           IF #Request AND NOT "PN_Mixinghead".Mixinghead[#MH].ReinigungskolbenDigital.ChckConnFault THEN
               "PN_Mixinghead".Mixinghead[#MH].ReinigungskolbenDigital.GeneralParameters.Request := "PN_Mixinghead".Mixinghead[#MH].ReinigungskolbenDigital.Active;
               "PN_Mixinghead".Mixinghead[#MH].ReinigungskolbenDigital.Zeiten.Request := "PN_Mixinghead".Mixinghead[#MH].ReinigungskolbenDigital.Active;
           END_IF;

           "WRREC_FC"(GOON := #GOON,
                      REQ := "PN_Mixinghead".Mixinghead[#MH].ReinigungskolbenDigital.GeneralParameters.Request,
                      ADDRESS := #TempHWID,
                      INDEX := #IDM_CleaningPiston_Digital_GeneralParameters_Index,
                      LENGTH := #IDM_CleaningPiston_Digital_GeneralParameters_Length,
                      WRREC_DONE => #t.DONE,
                      WRREC_BUSY => #t.BUSY,
                      WRREC_ERROR => #t.ERROR,
                      WRREC_STATUS => #t.STATUS,
                      ACTIVE := "PN_Mixinghead".Mixinghead[#MH].ReinigungskolbenDigital.Active,
                      RECORD := "PN_Mixinghead".Mixinghead[#MH].ReinigungskolbenDigital.GeneralParameters.Data,
                      DONE := "PN_Mixinghead".Mixinghead[#MH].ReinigungskolbenDigital.GeneralParameters.Transmitting);

           "WRREC_FC"(GOON := #GOON,
                      REQ := "PN_Mixinghead".Mixinghead[#MH].ReinigungskolbenDigital.Zeiten.Request,
                      ADDRESS := #TempHWID,
                      INDEX := #IDM_CleaningPiston_Digital_Zeiten_Index,
                      LENGTH := #IDM_CleaningPiston_Digital_Zeiten_Length,
                      WRREC_DONE => #t.DONE,
                      WRREC_BUSY => #t.BUSY,
                      WRREC_ERROR => #t.ERROR,
                      WRREC_STATUS => #t.STATUS,
                      ACTIVE := "PN_Mixinghead".Mixinghead[#MH].ReinigungskolbenDigital.Active,
                      RECORD := "PN_Mixinghead".Mixinghead[#MH].ReinigungskolbenDigital.Zeiten.Data,
                      DONE := "PN_Mixinghead".Mixinghead[#MH].ReinigungskolbenDigital.Zeiten.Transmitting);
       END_IF;

       // -----------------------------------
       // REINIGUNGSKOLBEN geregelt   
       // -----------------------------------
       IF "PN_Mixinghead".Mixinghead[#MH].ReinigungskolbenGeregelt.Active THEN
           #Address := INT_TO_WORD("PN_Mixinghead".Mixinghead[#MH].ReinigungskolbenGeregelt.Address);
           #ReturnValue := LOG2MOD(IOID := B#16#54, ADDR := #Address, HWID => #TempHWID);
           // Kommunikationsüberwachung
           // Nach einem Verbindungsabbruch werden die Telegramme automatisch verschickt.
           #Request := false;
           "CHCKPNCONN"(GOON := #GOON,
                        Active := "PN_Mixinghead".Mixinghead[#MH].ReinigungskolbenGeregelt.Active,
                        Address := #TempHWID,
                        PN_Request := #Request,
                        PN_Fault := "PN_Mixinghead".Mixinghead[#MH].ReinigungskolbenGeregelt.ChckConnFault,
                        DONE := "PN_Mixinghead".Mixinghead[#MH].ReinigungskolbenGeregelt.ChckConnDone);

           IF #Request AND NOT "PN_Mixinghead".Mixinghead[#MH].ReinigungskolbenGeregelt.ChckConnFault THEN
               "PN_Mixinghead".Mixinghead[#MH].ReinigungskolbenGeregelt.GeneralParameters.Request := "PN_Mixinghead".Mixinghead[#MH].ReinigungskolbenGeregelt.Active;
               "PN_Mixinghead".Mixinghead[#MH].ReinigungskolbenGeregelt.Zeiten.Request := "PN_Mixinghead".Mixinghead[#MH].ReinigungskolbenGeregelt.Active;
               "PN_Mixinghead".Mixinghead[#MH].ReinigungskolbenGeregelt.Skalierung.Request := "PN_Mixinghead".Mixinghead[#MH].ReinigungskolbenGeregelt.Active;
               "PN_Mixinghead".Mixinghead[#MH].ReinigungskolbenGeregelt.Regelparameter.Request := "PN_Mixinghead".Mixinghead[#MH].ReinigungskolbenGeregelt.Active;
           END_IF;

           "WRREC_FC"(GOON := #GOON,
                      REQ := "PN_Mixinghead".Mixinghead[#MH].ReinigungskolbenGeregelt.GeneralParameters.Request,
                      ACTIVE := "PN_Mixinghead".Mixinghead[#MH].ReinigungskolbenGeregelt.Active,
                      ADDRESS := #TempHWID,
                      INDEX := #IDM_CleaningPiston_Analog_Loop_GeneralParameters_Index,
                      LENGTH := #IDM_CleaningPiston_Analog_Loop_GeneralParameters_Length,
                      WRREC_DONE => #t.DONE,
                      WRREC_BUSY => #t.BUSY,
                      WRREC_ERROR => #t.ERROR,
                      WRREC_STATUS => #t.STATUS,
                      RECORD := "PN_Mixinghead".Mixinghead[#MH].ReinigungskolbenGeregelt.GeneralParameters.Data,
                      DONE := "PN_Mixinghead".Mixinghead[#MH].ReinigungskolbenGeregelt.GeneralParameters.Transmitting);

           "WRREC_FC"(GOON := #GOON,
                      REQ := "PN_Mixinghead".Mixinghead[#MH].ReinigungskolbenGeregelt.Zeiten.Request,
                      ACTIVE := "PN_Mixinghead".Mixinghead[#MH].ReinigungskolbenGeregelt.Active,
                      ADDRESS := #TempHWID,
                      INDEX := #IDM_CleaningPiston_Analog_Loop_Zeiten_Index,
                      LENGTH := #IDM_CleaningPiston_Analog_Loop_Zeiten_Length,
                      WRREC_DONE => #t.DONE,
                      WRREC_BUSY => #t.BUSY,
                      WRREC_ERROR => #t.ERROR,
                      WRREC_STATUS => #t.STATUS,
                      RECORD := "PN_Mixinghead".Mixinghead[#MH].ReinigungskolbenGeregelt.Zeiten.Data,
                      DONE := "PN_Mixinghead".Mixinghead[#MH].ReinigungskolbenGeregelt.Zeiten.Transmitting);

           "WRREC_FC"(GOON := #GOON,
                      REQ := "PN_Mixinghead".Mixinghead[#MH].ReinigungskolbenGeregelt.Skalierung.Request,
                      ACTIVE := "PN_Mixinghead".Mixinghead[#MH].ReinigungskolbenGeregelt.Active,
                      ADDRESS := #TempHWID,
                      INDEX := #IDM_Mixinghead_Digital_GeneralParameters_Index,
                      LENGTH := #IDM_Mixinghead_Digital_GeneralParameters_Length,
                      WRREC_DONE => #t.DONE,
                      WRREC_BUSY => #t.BUSY,
                      WRREC_ERROR => #t.ERROR,
                      WRREC_STATUS => #t.STATUS,
                      RECORD := "PN_Mixinghead".Mixinghead[#MH].ReinigungskolbenGeregelt.Skalierung.Data,
                      DONE := "PN_Mixinghead".Mixinghead[#MH].ReinigungskolbenGeregelt.Skalierung.Transmitting);

           "WRREC_FC"(GOON := #GOON,
                      REQ := "PN_Mixinghead".Mixinghead[#MH].ReinigungskolbenGeregelt.Regelparameter.Request,
                      ACTIVE := "PN_Mixinghead".Mixinghead[#MH].ReinigungskolbenGeregelt.Active,
                      ADDRESS := #TempHWID,
                      INDEX := #IDM_CleaningPiston_Analog_Loop_Regelparameter_Index,
                      LENGTH := #IDM_CleaningPiston_Analog_Loop_Regelparameter_Length,
                      WRREC_DONE => #t.DONE,
                      WRREC_BUSY => #t.BUSY,
                      WRREC_ERROR => #t.ERROR,
                      WRREC_STATUS => #t.STATUS,
                      RECORD := "PN_Mixinghead".Mixinghead[#MH].ReinigungskolbenGeregelt.Regelparameter.Data,
                      DONE := "PN_Mixinghead".Mixinghead[#MH].ReinigungskolbenGeregelt.Regelparameter.Transmitting);
       END_IF;

       // -----------------------------------
       // REINIGUNGSKOLBEN gesteuert   
       // -----------------------------------
       IF "PN_Mixinghead".Mixinghead[#MH].ReinigungskolbenGesteuert.Active THEN
           #Address := INT_TO_WORD("PN_Mixinghead".Mixinghead[#MH].ReinigungskolbenGesteuert.Address);
           #ReturnValue := LOG2MOD(IOID := B#16#54, ADDR := #Address, HWID => #TempHWID);
           // Kommunikationsüberwachung
           // Nach einem Verbindungsabbruch werden die Telegramme automatisch verschickt.
           #Request := false;
           "CHCKPNCONN"(GOON := #GOON,
                        Active := "PN_Mixinghead".Mixinghead[#MH].ReinigungskolbenGesteuert.Active,
                        Address := #TempHWID,
                        PN_Request := #Request,
                        PN_Fault := "PN_Mixinghead".Mixinghead[#MH].ReinigungskolbenGesteuert.ChckConnFault,
                        DONE := "PN_Mixinghead".Mixinghead[#MH].ReinigungskolbenGesteuert.ChckConnDone);

           IF #Request AND NOT "PN_Mixinghead".Mixinghead[#MH].ReinigungskolbenGesteuert.ChckConnFault THEN
               "PN_Mixinghead".Mixinghead[#MH].ReinigungskolbenGesteuert.GeneralParameters.Request := "PN_Mixinghead".Mixinghead[#MH].ReinigungskolbenGesteuert.Active;
               "PN_Mixinghead".Mixinghead[#MH].ReinigungskolbenGesteuert.Zeiten.Request := "PN_Mixinghead".Mixinghead[#MH].ReinigungskolbenGesteuert.Active;
               "PN_Mixinghead".Mixinghead[#MH].ReinigungskolbenGesteuert.Skalierung.Request := "PN_Mixinghead".Mixinghead[#MH].ReinigungskolbenGesteuert.Active;
               "PN_Mixinghead".Mixinghead[#MH].ReinigungskolbenGesteuert.StufenAktivierung.Request := "PN_Mixinghead".Mixinghead[#MH].ReinigungskolbenGesteuert.Active;
               "PN_Mixinghead".Mixinghead[#MH].ReinigungskolbenGesteuert.StufenRückkehr.Request := "PN_Mixinghead".Mixinghead[#MH].ReinigungskolbenGesteuert.Active;
           END_IF;

           "WRREC_FC"(GOON := #GOON,
                      REQ := "PN_Mixinghead".Mixinghead[#MH].ReinigungskolbenGesteuert.GeneralParameters.Request,
                      ACTIVE := "PN_Mixinghead".Mixinghead[#MH].ReinigungskolbenGesteuert.Active,
                      ADDRESS := #TempHWID,
                      INDEX := #IDM_CleaningPiston_Analog_GeneralParameters_Index,
                      LENGTH := #IDM_CleaningPiston_Analog_GeneralParameters_Length,
                      WRREC_DONE => #t.DONE,
                      WRREC_BUSY => #t.BUSY,
                      WRREC_ERROR => #t.ERROR,
                      WRREC_STATUS => #t.STATUS,
                      RECORD := "PN_Mixinghead".Mixinghead[#MH].ReinigungskolbenGesteuert.GeneralParameters.Data,
                      DONE := "PN_Mixinghead".Mixinghead[#MH].ReinigungskolbenGesteuert.GeneralParameters.Transmitting);

           "WRREC_FC"(GOON := #GOON,
                      REQ := "PN_Mixinghead".Mixinghead[#MH].ReinigungskolbenGesteuert.Zeiten.Request,
                      ACTIVE := "PN_Mixinghead".Mixinghead[#MH].ReinigungskolbenGesteuert.Active,
                      ADDRESS := #TempHWID,
                      INDEX := #IDM_CleaningPiston_Analog_Zeiten_Index,
                      LENGTH := #IDM_CleaningPiston_Analog_Zeiten_Length,
                      WRREC_DONE => #t.DONE,
                      WRREC_BUSY => #t.BUSY,
                      WRREC_ERROR => #t.ERROR,
                      WRREC_STATUS => #t.STATUS,
                      RECORD := "PN_Mixinghead".Mixinghead[#MH].ReinigungskolbenGesteuert.Zeiten.Data,
                      DONE := "PN_Mixinghead".Mixinghead[#MH].ReinigungskolbenGesteuert.Zeiten.Transmitting);

           "WRREC_FC"(GOON := #GOON,
                      REQ := "PN_Mixinghead".Mixinghead[#MH].ReinigungskolbenGesteuert.Skalierung.Request,
                      ACTIVE := "PN_Mixinghead".Mixinghead[#MH].ReinigungskolbenGesteuert.Active,
                      ADDRESS := #TempHWID,
                      INDEX := #IDM_CleaningPiston_Analog_Skalierung_Index,
                      LENGTH := #IDM_CleaningPiston_Analog_Skalierung_Length,
                      WRREC_DONE => #t.DONE,
                      WRREC_BUSY => #t.BUSY,
                      WRREC_ERROR => #t.ERROR,
                      WRREC_STATUS => #t.STATUS,
                      RECORD := "PN_Mixinghead".Mixinghead[#MH].ReinigungskolbenGesteuert.Skalierung.Data,
                      DONE := "PN_Mixinghead".Mixinghead[#MH].ReinigungskolbenGesteuert.Skalierung.Transmitting);

           "WRREC_FC"(GOON := #GOON,
                      REQ := "PN_Mixinghead".Mixinghead[#MH].ReinigungskolbenGesteuert.StufenAktivierung.Request,
                      ACTIVE := "PN_Mixinghead".Mixinghead[#MH].ReinigungskolbenGesteuert.Active,
                      ADDRESS := #TempHWID,
                      INDEX := #IDM_CleaningPiston_Analog_StufenAktivierung_Index,
                      LENGTH := #IDM_CleaningPiston_Analog_StufenAktivierung_Length,
                      WRREC_DONE => #t.DONE,
                      WRREC_BUSY => #t.BUSY,
                      WRREC_ERROR => #t.ERROR,
                      WRREC_STATUS => #t.STATUS,
                      RECORD := "PN_Mixinghead".Mixinghead[#MH].ReinigungskolbenGesteuert.StufenAktivierung.Data,
                      DONE := "PN_Mixinghead".Mixinghead[#MH].ReinigungskolbenGesteuert.StufenAktivierung.Transmitting);

           "WRREC_FC"(GOON := #GOON,
                      REQ := "PN_Mixinghead".Mixinghead[#MH].ReinigungskolbenGesteuert.StufenRückkehr.Request,
                      ACTIVE := "PN_Mixinghead".Mixinghead[#MH].ReinigungskolbenGesteuert.Active,
                      ADDRESS := #TempHWID,
                      INDEX := #IDM_CleaningPiston_Analog_StufenRückkehr_Index,
                      LENGTH := #IDM_CleaningPiston_Analog_StufenRückkehr_Length,
                      WRREC_DONE => #t.DONE,
                      WRREC_BUSY => #t.BUSY,
                      WRREC_ERROR => #t.ERROR,
                      WRREC_STATUS => #t.STATUS,
                      RECORD := "PN_Mixinghead".Mixinghead[#MH].ReinigungskolbenGesteuert.StufenRückkehr.Data,
                      DONE := "PN_Mixinghead".Mixinghead[#MH].ReinigungskolbenGesteuert.StufenRückkehr.Transmitting);
       END_IF;

       // -----------------------------------
       // Düse/Bypass   
       // -----------------------------------
       FOR #DB := 1 TO 8 DO
           IF "PN_Mixinghead".Mixinghead[#MH].DüseBypass[#DB].Active THEN
               #Address := INT_TO_WORD("PN_Mixinghead".Mixinghead[#MH].DüseBypass[#DB].Address);
               #ReturnValue := LOG2MOD(IOID := B#16#54, ADDR := #Address, HWID => #TempHWID);
               // Kommunikationsüberwachung
               // Nach einem Verbindungsabbruch werden die Telegramme automatisch verschickt.
               #Request := false;
               "CHCKPNCONN"(GOON := #GOON,
                            Active := "PN_Mixinghead".Mixinghead[#MH].DüseBypass[#DB].Active,
                            Address := #TempHWID,
                            PN_Request := #Request,
                            PN_Fault := "PN_Mixinghead".Mixinghead[#MH].DüseBypass[#DB].ChckConnFault,
                            DONE := "PN_Mixinghead".Mixinghead[#MH].DüseBypass[#DB].ChckConnDone);

               IF #Request AND NOT "PN_Mixinghead".Mixinghead[#MH].DüseBypass[#DB].ChckConnFault THEN
                   "PN_Mixinghead".Mixinghead[#MH].DüseBypass[#DB].Zeiten.Request := "PN_Mixinghead".Mixinghead[#MH].DüseBypass[#DB].Active;
               END_IF;

               "WRREC_FC"(GOON := #GOON,
                          REQ := "PN_Mixinghead".Mixinghead[#MH].DüseBypass[#DB].Zeiten.Request,
                          ACTIVE := "PN_Mixinghead".Mixinghead[#MH].DüseBypass[#DB].Active,
                          ADDRESS := #TempHWID,
                          INDEX := #IDM_Mixinghead_NozzleBypass_Zeiten_Index,
                          LENGTH := #IDM_Mixinghead_NozzleBypass_Zeiten_Length,
                          WRREC_DONE => #t.DONE,
                          WRREC_BUSY => #t.BUSY,
                          WRREC_ERROR => #t.ERROR,
                          WRREC_STATUS => #t.STATUS,
                          RECORD := "PN_Mixinghead".Mixinghead[#MH].DüseBypass[#DB].Zeiten.Data,
                          DONE := "PN_Mixinghead".Mixinghead[#MH].DüseBypass[#DB].Zeiten.Transmitting);
           END_IF;
       END_FOR;
   END_FOR;
END_FUNCTION

FUNCTION "WRREC_FC" : Void   // FC1007, SCL
{ S7_Optimized_Access := 'FALSE' }
VERSION : 0.1
   VAR_INPUT
      ADDRESS : Hw_Io;   // Adresse des zu parametrierenden IO-Bereichs
      INDEX : Int;   // Index des zu sendenden Telegrams
      LENGTH : Int;   // Länge des zu sendenden Telegrams
   END_VAR
   VAR_OUTPUT
      WRREC_DONE : Bool;   // Datensatz wurde übertragen
      WRREC_BUSY : Bool;   // Schreibvorgang ist noch nicht beendet
      WRREC_ERROR : Bool;   // Fehler beim Schreibvorgang
      WRREC_STATUS : DWord;   // Bausteinstatus und Fehlerinformation
   END_VAR
   VAR_IN_OUT
      GOON : Bool;
      REQ : Bool;   // Anforderung zum Datenaustausch
      ACTIVE : Bool;   // Generelle Freigabe Datenübertragung
      RECORD : ANY;   // Datensatz
      DONE : Bool;   // Zeigt an, dass die Übertragung für diesen Aufruf gestartet wurde.
   END_VAR
   VAR_TEMP
      i : Int;
   END_VAR
BEGIN
   // Der Baustein WRREC_FC überträgt Telegramme an Profinetteilnehmer,
   // um Parameter zu ändern. Anpassungen in der Hardwarekonfiguration
   // sind damit nicht notwendig. Somit entfällt auch die Übersetzung,
   // Übertragung der Hardwarekonfiguration und der Neustart der CPU.
   // 
   // Der IOs dieses FCs ist nahezu identisch zu WRREC. Die Bedeutung der
   // Variablen kann also in der Hilfe nachgelesen werden.
   // Zweck dieses Bausteins ist es, alle Telegramme über einen WRREC-Aufruf
   // zu verschicken. So ist nur ein Instanz-DB nötig.

   // =======================================================================
   // 
   // Bearbeite die Funktion, wenn die Funktion eine Übertragung gestartet oder,
   // wenn keine Übertragung stattfindet

   IF NOT #GOON THEN
       #DONE := false;
   END_IF;

   IF #ACTIVE THEN
       IF #GOON AND NOT #DONE THEN
           "WRREC_DB"(REQ := #REQ,
                      ID := #ADDRESS,
                      INDEX := #INDEX,
                      LEN := INT_TO_UINT(#LENGTH),
                      DONE => #WRREC_DONE,
                      BUSY => #WRREC_BUSY,
                      ERROR => #WRREC_ERROR,
                      STATUS => #WRREC_STATUS,
                      RECORD := #RECORD);

           IF (#WRREC_BUSY = 0) OR #WRREC_DONE OR #WRREC_ERROR THEN
               // Bearbeitung beendet
               #DONE := true;
               // Request setzen, wenn ein Fehler ermittelt wurde. 
               #REQ := #WRREC_ERROR;
           END_IF;
           // Fehler ausgeben
           IF #WRREC_ERROR THEN
               // Sammelstörung setzen und Meldung ausgeben.
               // 
               "PN_Error".Fault := true;
               // Index 1 enthält immer die aktuellste Meldung. Bei einer neuen Meldung
               // werden alle anderen ein Arrayelement weitergeschoben.
               // 
               FOR #i := 9 TO 1 BY -1 DO
                   "PN_Error".Error[#i + 1].Address := "PN_Error".Error[#i].Address;
                   "PN_Error".Error[#i + 1].Index := "PN_Error".Error[#i].Index;
                   "PN_Error".Error[#i + 1].Length := "PN_Error".Error[#i].Length;
                   "PN_Error".Error[#i + 1].State := "PN_Error".Error[#i].State;
               END_FOR;

               "PN_Error".Error[1].Address := #ADDRESS;
               "PN_Error".Error[1].Index := #INDEX;
               "PN_Error".Error[1].Length := #LENGTH;
               "PN_Error".Error[1].State := #WRREC_STATUS;
           END_IF;
       END_IF;
   ELSE
       #DONE := #GOON;
   END_IF;

   #GOON := #DONE;

   // Reset setzt alle Fehlerausgaben zurück.
   // 
   IF "PN_Error".Reset THEN
       FOR #i := 1 TO 10 DO
           "PN_Error".Error[#i].Address := 0;
           "PN_Error".Error[#i].Index := 0;
           "PN_Error".Error[#i].Length := 0;
           "PN_Error".Error[#i].State := 0;
           "PN_Error".Reset := false;
       END_FOR;
   END_IF;




   // ALTER CODE
   // IF #TRANSMITTING OR ((NOT "WRREC_DB".BUSY) AND #ACTIVE) THEN
   //     "WRREC_DB"(REQ := #REQ,
   //                  ID := #ADDRESS,
   //                  INDEX := #INDEX,
   //                  LEN := #LENGTH,
   //                  DONE => #WRREC_DONE,
   //                  BUSY => #WRREC_BUSY,
   //                  ERROR => #WRREC_ERROR,
   //                  STATUS => #WRREC_STATUS,
   //                  RECORD := #RECORD);

   //     // Setze REQ zurück, wenn Übertragung beendet ist
   //       IF #WRREC_DONE THEN
   //           #REQ := false;
   //       END_IF;

   //       #TRANSMITTING := #REQ AND NOT (#WRREC_DONE OR #WRREC_ERROR);

   //     IF #WRREC_ERROR THEN
   //         // Sammelstörung setzen und Meldung ausgeben.
   //         // 
   //         "PN_Error".Fault := true;
   //         // Index 1 enthält immer die aktuellste Meldung. Bei einer neuen Meldung
   //         // werden alle anderen ein Arrayelement weitergeschoben.
   //         // 
   //         FOR #i := 9 TO 1 BY -1 DO
   //             "PN_Error".Error[#i + 1].Address := "PN_Error".Error[#i].Address;
   //             "PN_Error".Error[#i + 1].Index := "PN_Error".Error[#i].Index;
   //             "PN_Error".Error[#i + 1].Length := "PN_Error".Error[#i].Length;
   //             "PN_Error".Error[#i + 1].State := "PN_Error".Error[#i].State;
   //         END_FOR;

   //         "PN_Error".Error[1].Address := #ADDRESS;
   //         "PN_Error".Error[1].Index := #INDEX;
   //         "PN_Error".Error[1].Length := #LENGTH;
   //         "PN_Error".Error[1].State := #WRREC_STATUS;
   //     END_IF;
   // END_IF;
   // // Reset setzt alle Fehlerausgaben zurück.
   // // 
   // IF "PN_Error".Reset THEN
   //     FOR #i := 1 TO 10 DO
   //         "PN_Error".Error[#i].Address := 0;
   //         "PN_Error".Error[#i].Index := 0;
   //         "PN_Error".Error[#i].Length := 0;
   //         "PN_Error".Error[#i].State := 0;
   //         "PN_Error".Reset := false;
   //     END_FOR;
   // END_IF;
END_FUNCTION

FUNCTION "FC1001_TT" : Void   // FC1010, STL
TITLE = Dryside Turntable and additional devices
{ S7_Optimized_Access := 'TRUE' }
VERSION : 0.1
BEGIN

REGION Network 1
         CALL  "FC1011_TT_Fault";
         CALL  "FC1021_TT_Operation_mode";
         CALL  "FC1031_AdditionalDevice";
         CALL  "FC1040_TT_Movement";
         CALL  "FC1051_TT_Segment";
END_REGION
END_FUNCTION

FUNCTION "FC1011_TT_Fault" : Void   // FC1011, STL
{ S7_Optimized_Access := 'TRUE' }
VERSION : 0.1
   VAR_TEMP
      Dummy_Bit_fuer_PUC : Bool;
   END_VAR
BEGIN

REGION Network 1: Bit zum Zurücksetzen der Störungen in den einzelnen FC`s Rundtisch 1
         A     "DB009_Faults".Faults_Reset_FKT_M1;
         =     "DB1011_TT_Fault".Reset_FC_RT;
         A     "DB009_Faults".Faults_Reset_Group;
         =     "DB1011_TT_Fault".Reset_STGR_RT;
END_REGION

REGION Network 2
   //-----
         CALL  "FC1012_TT_Fault"
         ( IN_Reset_fault_Grp      := "DB1011_TT_Fault".Reset_STGR_RT,
           IN_TT_Exist             := "DB1009_TT_Config".Bit.WithTT,
           IN_Erster_SPS_Zyklus    := "FirstScan",
           IN_Stoer_Grp_1_von_Ext  := FALSE,
           IN_Stoer_Grp_2_von_Ext  := FALSE,
           IN_Stoer_Grp_3_von_Ext  := FALSE,
           IN_DB_Stoerungen        := "DB1011_TT_Fault",
           IN_Start_Stoerungen     := 2,
           IO_Stoer_Grp_1_aktiv    := "DB1011_TT_Fault".STG1_RT,
           IO_Stoer_Grp_2_aktiv    := "DB1011_TT_Fault".STG2_RT,
           IO_Stoer_Grp_3_aktiv    := "DB1011_TT_Fault".STG3_RT,
           IO_Stoerungsaenderung   := "DB1011_TT_Fault".Stoerungsaend_RT,
           IO_FM_Stoer_Grp_1_v_Ext := "DB1011_TT_Fault".FHM_NeuStoer_Grp_1,
           IO_FM_Stoer_Grp_2_v_Ext := "DB1011_TT_Fault".FHM_NeuStoer_Grp_2,
           IO_FM_Stoer_Grp_3_v_Ext := "DB1011_TT_Fault".FHM_NeuStoer_Grp_3,
           IO_Daten_Senden         := #Dummy_Bit_fuer_PUC
         );
   //-----
END_REGION

REGION Network 3: A fault exist at the dryside
         O     "DB1011_TT_Fault".STG1_RT;
         O     "DB1011_TT_Fault".STG2_RT;
         O     "DB1011_TT_Fault".STG3_RT;
         =     "DB1001_TT_State".Bits.Fault_Exist;
END_REGION

REGION Network 4: In der Steuerung wurde eine Störung der Gruppe 1 der Fremdanlage festgestellt
         A     "DB1011_TT_Fault".STG1_RT;
         =     "DB009_Faults".Faults_FKT_Grp_1_ExtP;
         A     "DB1011_TT_Fault".STG2_RT;
         =     "DB009_Faults".Faults_FKT_Grp_2_ExtP;
         A     "DB1011_TT_Fault".STG3_RT;
         =     "DB009_Faults".Faults_FKT_Grp_3_ExtP;
         A     "DB1011_TT_Fault".Stoerungsaend_RT;
         S     "DB009_Faults".Faultschanging_ExtP;
         R     "DB1011_TT_Fault".Stoerungsaend_RT;
END_REGION
END_FUNCTION

FUNCTION "FC1012_TT_Fault" : Void   // FC1012, STL
TITLE = Stoerungsgruppe 1
{ S7_Optimized_Access := 'FALSE' }
AUTHOR : KT242
VERSION : 0.1
   VAR_INPUT
      IN_Reset_fault_Grp : Bool;   // Signal zum ablöschen der Störungen innerhalb des Störungsbausteins
      IN_TT_Exist : Bool;   // Selection that a turntable exist
      IN_Erster_SPS_Zyklus : Bool;   // Impulssignal Neusstart der Steuerung zum ablöschen der Störungen
      IN_Stoer_Grp_1_von_Ext : Bool;   // Eine Störung der Gruppe 1 vom Extern (zB. übergeordente Funktion) steht an
      IN_Stoer_Grp_2_von_Ext : Bool;   // Eine Störung der Gruppe 2 vom Extern (zB. übergeordente Funktion) steht an
      IN_Stoer_Grp_3_von_Ext : Bool;   // Eine Störung der Gruppe 3 vom Extern (zB. übergeordente Funktion) steht an
      IN_DB_Stoerungen : DB_ANY;   // Nummer des Datenbausteins zum "Zwischenmerken" der Störungen
      IN_Start_Stoerungen : Int;   // Startadresse der Störungen im Störungsbaustein für diese Maschine
   END_VAR
   VAR_IN_OUT
      IO_Stoer_Grp_1_aktiv : Bool;   // An diesem Formträger steht eine Störung der Gruppe 1 an
      IO_Stoer_Grp_2_aktiv : Bool;   // An diesem Formträger steht eine Störung der Gruppe 2 an
      IO_Stoer_Grp_3_aktiv : Bool;   // An diesem Formträger steht eine Störung der Gruppe 3 an
      IO_Stoerungsaenderung : Bool;   // Eine eingehende neue Störung wurde erkannt
      IO_FM_Stoer_Grp_1_v_Ext : Bool;   // Flankenmerker für die Erkennung einer neuen Störung der Gruppe 1 von Extern
      IO_FM_Stoer_Grp_2_v_Ext : Bool;   // Flankenmerker für die Erkennung einer neuen Störung der Gruppe 2 von Extern
      IO_FM_Stoer_Grp_3_v_Ext : Bool;   // Flankenmerker für die Erkennung einer neuen Störung der Gruppe 3 von Extern
      IO_Daten_Senden : Bool;   // Signal für die Übertragung der Störungen eine übergeordnete SPS
   END_VAR
   VAR_TEMP
      St_Nr_009 : Bool;
      St_Nr_010 : Bool;
      St_Nr_011 : Bool;
      St_Nr_012 : Bool;
      St_Nr_013 : Bool;
      St_Nr_014 : Bool;
      St_Nr_015 : Bool;
      St_Nr_016 : Bool;
      St_Nr_001 : Bool;
      St_Nr_002 : Bool;
      St_Nr_003 : Bool;
      St_Nr_004 : Bool;
      St_Nr_005 : Bool;
      St_Nr_006 : Bool;
      St_Nr_007 : Bool;
      St_Nr_008 : Bool;
      St_Nr_025 : Bool;
      St_Nr_026 : Bool;
      St_Nr_027 : Bool;
      St_Nr_028 : Bool;
      St_Nr_029 : Bool;
      St_Nr_030 : Bool;
      St_Nr_031 : Bool;
      St_Nr_032 : Bool;
      St_Nr_017 : Bool;
      St_Nr_018 : Bool;
      St_Nr_019 : Bool;
      St_Nr_020 : Bool;
      St_Nr_021 : Bool;
      St_Nr_022 : Bool;
      St_Nr_023 : Bool;
      St_Nr_024 : Bool;
      St_Nr_041 : Bool;
      St_Nr_042 : Bool;
      St_Nr_043 : Bool;
      St_Nr_044 : Bool;
      St_Nr_045 : Bool;
      St_Nr_046 : Bool;
      St_Nr_047 : Bool;
      St_Nr_048 : Bool;
      St_Nr_033 : Bool;
      St_Nr_034 : Bool;
      St_Nr_035 : Bool;
      St_Nr_036 : Bool;
      St_Nr_037 : Bool;
      St_Nr_038 : Bool;
      St_Nr_039 : Bool;
      St_Nr_040 : Bool;
      St_Nr_057 : Bool;
      St_Nr_058 : Bool;
      St_Nr_059 : Bool;
      St_Nr_060 : Bool;
      St_Nr_061 : Bool;
      St_Nr_062 : Bool;
      St_Nr_063 : Bool;
      St_Nr_064 : Bool;
      St_Nr_049 : Bool;
      St_Nr_050 : Bool;
      St_Nr_051 : Bool;
      St_Nr_052 : Bool;
      St_Nr_053 : Bool;
      St_Nr_054 : Bool;
      St_Nr_055 : Bool;
      St_Nr_056 : Bool;
      St_Nr_073 : Bool;
      St_Nr_074 : Bool;
      St_Nr_075 : Bool;
      St_Nr_076 : Bool;
      St_Nr_077 : Bool;
      St_Nr_078 : Bool;
      St_Nr_079 : Bool;
      St_Nr_080 : Bool;
      St_Nr_065 : Bool;
      St_Nr_066 : Bool;
      St_Nr_067 : Bool;
      St_Nr_068 : Bool;
      St_Nr_069 : Bool;
      St_Nr_070 : Bool;
      St_Nr_071 : Bool;
      St_Nr_072 : Bool;
      St_Nr_089 : Bool;
      St_Nr_090 : Bool;
      St_Nr_091 : Bool;
      St_Nr_092 : Bool;
      St_Nr_093 : Bool;
      St_Nr_094 : Bool;
      St_Nr_095 : Bool;
      St_Nr_096 : Bool;
      St_Nr_081 : Bool;
      St_Nr_082 : Bool;
      St_Nr_083 : Bool;
      St_Nr_084 : Bool;
      St_Nr_085 : Bool;
      St_Nr_086 : Bool;
      St_Nr_087 : Bool;
      St_Nr_088 : Bool;
      Mld_Nr_105 : Bool;
      Mld_Nr_106 : Bool;
      Mld_Nr_107 : Bool;
      Mld_Nr_108 : Bool;
      Mld_Nr_109 : Bool;
      Mld_Nr_110 : Bool;
      Mld_Nr_111 : Bool;
      Mld_Nr_112 : Bool;
      Mld_Nr_097 : Bool;
      Mld_Nr_098 : Bool;
      Mld_Nr_099 : Bool;
      Mld_Nr_100 : Bool;
      Mld_Nr_101 : Bool;
      Mld_Nr_102 : Bool;
      Mld_Nr_103 : Bool;
      Mld_Nr_104 : Bool;
      Mld_Nr_121 : Bool;
      Mld_Nr_122 : Bool;
      Mld_Nr_123 : Bool;
      Mld_Nr_124 : Bool;
      Mld_Nr_125 : Bool;
      Mld_Nr_126 : Bool;
      Mld_Nr_127 : Bool;
      Mld_Nr_128 : Bool;
      Mld_Nr_113 : Bool;
      Mld_Nr_114 : Bool;
      Mld_Nr_115 : Bool;
      Mld_Nr_116 : Bool;
      Mld_Nr_117 : Bool;
      Mld_Nr_118 : Bool;
      Mld_Nr_119 : Bool;
      Mld_Nr_120 : Bool;
      Schleifenzaehler : Int;
   END_VAR
BEGIN

REGION Network 1: Stoerungen auf Lokaldaten schreiben oder quittieren
   // Wenn aus dem Quittierungsbaustein (FB9; FC9) das Bit zum ablöschen der 
   // Störungen gesetzt wird (2´tes mal quittiert) werden die lokalen Störungen der 
   // Gruppe 1 bis 3 abgelöscht.
   // Ansonsten werden die im Datenbaustein gespeicherten Störungen auf die Lokalen 
   // übertragen.
         O     #IO_Stoer_Grp_1_aktiv;  // Wenn eine Sammelstörung der drei
         O     #IO_Stoer_Grp_2_aktiv;  // Störunggruppen noch ansteht,
         O     #IO_Stoer_Grp_3_aktiv;  // und die Quittierung erfolgt oder
         A     #IN_Reset_fault_Grp;  // beim Neustart der Steuerung werden die
         O     #IN_Erster_SPS_Zyklus;  // Sammelstörungen der Gruppen abgelöscht
         ON    #IN_TT_Exist;
         R     #IO_Stoer_Grp_1_aktiv;  // und die Sendeanforderung gesetzt.
         R     #IO_Stoer_Grp_2_aktiv;  // Dieses muß erfolgen, da sonst die letzte
         R     #IO_Stoer_Grp_3_aktiv;  // angezeigte Störung nicht in der Visualisierung
         S     #IO_Daten_Senden;  // ausgetragen wird.
   //
         L     0;  // Interner Offset für Störungsgruppe 1
         SLD   3;  //
         LAR1;  // Adresse für lokale Störungen
   //
         L     0;  // Interner Offset für Störungsgruppe 1
         L     #IN_Start_Stoerungen;
         +D;
         SLD   3;  //
         LAR2;  // Adresse für Störung im DB
   //
         L     6;  // Anzahl der Störungsworte
   M001: T     #Schleifenzaehler;  // Störungsgruppe 1+ 2 +3
         OPN   #IN_DB_Stoerungen;  // Öffnen des Störungsbausteins
         L     DBW[AR2, P#0.0];  // Gespeicherte Störung auf lokale schreiben
         A     #IN_Reset_fault_Grp;  // Bei Quittierung werden die
         JCN   M002;  // Störungen zurückgesetzt
         L     0;  //
         T     DBW[AR2, P#0.0];  // die gespeicherten und die
   M002: T     LW[AR1, P#0.0];  // Lokalen Störungen
   //
         +AR1  P#2.0;
         +AR2  P#2.0;
   //
         L     #Schleifenzaehler;  // Wenn Schleifenzähler <> 0
         LOOP  M001;  // Schleife erneut durchlaufen
   //
         AN    #IN_TT_Exist;
         BEU;
END_REGION

REGION Network 2: Störungsbits Störungen Gruppe 1
   // am OP ab 81 !
         NOP   0;
   // 001 SEW-Umrichter für Rundtischantrieb am Profibus nicht erreichbar
         A     "DB1040_TT_MovementFault".IPOS.STG_Busfehler;
         S     #St_Nr_001;
   // 002 Störung Segmentkennung: Nummer unlogisch
         A     "DB1040_TT_MovementFault".Segmentkennung.STG_Nummer_unlogisch;
         S     #St_Nr_002;
   // 003 Zentrale am Profibs nihct erreichbar
   //    U     "Flag_DP_Bus1_ADR007_ok"
   //    S     #St_Nr_003
   // 004 Dezentrale auf Rundtisch am Profibus nicht erreichbar
   //    S     #St_Nr_004
   // 005 Anlagenbetrieb stoppen
   //     S     #St_Nr_005
   // 006 Schäummaschine oder Roboter nicht bereit
   //     S     #St_Nr_006
   // 007 Umrichter Rundtischantrieb nicht betriebsbereit
         A     "DB1040_TT_MovementFault".IPOS.STG_Umrichter;
         S     #St_Nr_007;
   // 008 Störung Motorschutz Rundtischantrieb
         A     "DB1040_TT_MovementFault".IPOS.STG_Motorschutz;
         S     #St_Nr_008;
   // 009 Störung SEW Umrichter RT Antrieb
         O     "DB1040_TT_MovementFault".IPOS.STG_von_IPOS;
         S     #St_Nr_009;
   // 010 Störung Genauhaltini
   //      U     "DB151_Rundtisch_1".IPOS.Status.RT_dreht
   //      FP    "FHM_RT1_dreht"
   //      =     "HM_RT1_dreht"
   //
   //      O     "HM_RT1_dreht"
   //      O     "DB009_Stoerungen".Reset_FC_RT_01
   //      R     "HM_RT1_Ziel_erreicht"
   //
   //      U     "DB151_Rundtisch_1".IPOS.Eingaenge_von_IPOS.Ziel_erreicht
   //      U     "DB151_Rundtisch_1".IPOS.Status.IPOS_referenziert
   //      S     "HM_RT1_Ziel_erreicht"
   //
   //      U     "HM_RT1_Ziel_erreicht"
   //      U     "DB151_Rundtisch_1".BA_Anlage.Produktion
   //      UN    "DB151_Rundtisch_1".BA_Anlage.Referenzieren
   //      UN    "GenauhaltINI"
   //      L     S5T#3S
   //      SE    "Tag_19"
   //
   //      U     "Tag_19"
   //      CLR
   //      S     #St_Nr_010
   // 011 Es ist keine Segmentkennung vorhanden
         A     "DB1050_Seg_Fault".Segmentverwaltung.STG_keine_SegmentNr;
         S     #St_Nr_011;
   // 012 Das Paritätsbit wurde falsch gesetzt
         A     "DB1050_Seg_Fault".Segmentverwaltung.STG_falsche_Paritaet;
         S     #St_Nr_012;
   // 013 Die verdrahtete Segmentnummer ist für dieses RT zu groß
         A     "DB1050_Seg_Fault".Segmentverwaltung.STG_SegNr_zu_gross;
         S     #St_Nr_013;
   // 014 Der Platz auf dem Segment wurde doppelt belegt // Verdrahtungsfehler
         A     "DB1050_Seg_Fault".Segmentverwaltung.STG_Platz_doppelt;
         S     #St_Nr_014;
   // 015 Formnummer wechselt im laufenden Betrieb
   //       O     "DB201_RT1_Segment_1".Status_FT.Segment_Bits.STG_Nummer_wechselt
   //       O     "DB202_RT1_Segment_2".Status_FT.Segment_Bits.STG_Nummer_wechselt
   //       O     "DB203_RT1_Segment_3".Status_FT.Segment_Bits.STG_Nummer_wechselt
   //       O     "DB204_RT1_Segment_4".Status_FT.Segment_Bits.STG_Nummer_wechselt
   //       O     "DB205_RT1_Segment_5".Status_FT.Segment_Bits.STG_Nummer_wechselt
   //       O     "DB206_RT1_Segment_6".Status_FT.Segment_Bits.STG_Nummer_wechselt
   //       O     "DB207_RT1_Segment_7".Status_FT.Segment_Bits.STG_Nummer_wechselt
   //       O     "DB208_RT1_Segment_8".Status_FT.Segment_Bits.STG_Nummer_wechselt
   //       O     "DB209_RT1_Segment_9".Status_FT.Segment_Bits.STG_Nummer_wechselt
   //       O     "DB210_RT1_Segment_10".Status_FT.Segment_Bits.STG_Nummer_wechselt
   //       O     "DB211_RT1_Segment_11".Status_FT.Segment_Bits.STG_Nummer_wechselt
   //       O     "DB213_RT1_Segment_13".Status_FT.Segment_Bits.STG_Nummer_wechselt
   //       O     "DB214_RT1_Segment_14".Status_FT.Segment_Bits.STG_Nummer_wechselt
   //       O     "DB215_RT1_Segment_15".Status_FT.Segment_Bits.STG_Nummer_wechselt
   //       O     "DB216_RT1_Segment_16".Status_FT.Segment_Bits.STG_Nummer_wechselt
   //       O     "DB217_RT1_Segment_17".Status_FT.Segment_Bits.STG_Nummer_wechselt
   //       O     "DB218_RT1_Segment_18".Status_FT.Segment_Bits.STG_Nummer_wechselt
   //       O     "DB219_RT1_Segment_19".Status_FT.Segment_Bits.STG_Nummer_wechselt
   //       O     "DB220_RT1_Segment_20".Status_FT.Segment_Bits.STG_Nummer_wechselt
   //       S     #St_Nr_015

   // 016 Störung von IPOS
         A     "DB1040_TT_MovementFault".IPOS.STG_von_IPOS;
         S     #St_Nr_016;
   // 017 Störung Segmentkennung: falsche Hardwareabschaltung
         A     "DB1040_TT_MovementFault".Segmentkennung.STG_Hardwareabschaltung;
         S     #St_Nr_017;
   // 018 Genauhaltini defekt oder immer bedeckt
         A     "DB1040_TT_MovementFault".IPOS.STG_Genauhalt_immer_ein;
         S     #St_Nr_018;
   // 019 Reserve
   //      S     #St_Nr_019
   // 020 Reserve
   //    S     #St_Nr_020
   // 021 Reserve
   //    S     #St_Nr_021
   // 022 Reserve
   //    S     #St_Nr_022
   // 023 Reserve
   //    S     #St_Nr_023
   // 024 Reserve
   //    S     #St_Nr_024
   // 025 Reserve
   //    S     #St_Nr_025
   // 026 Reserve
   //    S     #St_Nr_026
   // 027 Reserve
   //    S     #St_Nr_027
   // 028 Reserve
   //    S     #St_Nr_028
   // 029 Reserve
   //    S     #St_Nr_029
   // 030 Reserve
   //    S     #St_Nr_030
   // 031 Reserve
   //    S     #St_Nr_031
   // 032 Reserve
   //    S     #St_Nr_032
END_REGION

REGION Network 3: Stoerungsbits Störungen Gruppe 2
         NOP   0;
   // 033 Störung Lüfter Umrichter Rundtischantrieb
         A     "DB1040_TT_MovementFault".IPOS.STG_Luefter;
         S     #St_Nr_033;
   // 034 Reserve
   //    S     #St_Nr_034
   // 035 Reserve
   //    S     #St_Nr_035
   // 036 Reserve
   //    S     #St_Nr_036
   // 037 Reserve
   //    S     #St_Nr_037
   // 038 Reserve
   //    S     #St_Nr_038
   // 039 Reserve
   //    S     #St_Nr_039
   // 040 Reserve
   //    S     #St_Nr_040
   // 041 Reserve
   //    S     #St_Nr_041
   // 042 Reserve
   //    S     #St_Nr_042
   // 043 Reserve
   //    S     #St_Nr_043
   // 044 Reserve
   //    S     #St_Nr_044
   // 045 Reserve
   //    S     #St_Nr_045
   // 046 Reserve
   //    S     #St_Nr_046
   // 047 Reserve
   //    S     #St_Nr_047
   // 048 Reserve
   //    S     #St_Nr_048
END_REGION

REGION Network 4: Stoerungsbits Störungen Gruppe 3
         NOP   0;
   // 049 Störung Sicherung Segmente
   //      S     #St_Nr_049
   // 050 Störung Versorgung Bremse des Rundtisches
   //       UN    "F_Bremse_RT_1"
   //       S     #St_Nr_050
   // 051 Eine Sicherheitseinrichtung für Tippbetrieb nicht quittiert
         O     "Button_Tip_+";
         O     "Button_Tip_-";
         A     "DB1001_TT_State".BA_Anlage.Hand;
         A(;
         O     "DB1031_AddStatus".SaftyDevice[1].HFforMESAutomaticStop;
         O     "DB1031_AddStatus".SaftyDevice[2].HFforMESAutomaticStop;
         O     "DB1031_AddStatus".SaftyDevice[3].HFforMESAutomaticStop;
         O     "DB1031_AddStatus".SaftyDevice[4].HFforMESAutomaticStop;
         ON    "AS_pendelum_flap_to_handling";
         ON    "AS_pendelum_flap_from_handling";
         );
         S     #St_Nr_051;
   // 052 Störung Versorgung Schleifring
   //    S     #St_Nr_052
   // 053 Schäumroboter nicht bereit
   //    U     "T_Start_RT_1"
   //    U     "DB151_Rundtisch_1".BA_Anlage.Automatik
   //    UN    "DB005_RS<->Extern".Status_RS.Frg_Roboter_f_Schaeumen
   //    U     "DB005_RS<->Extern".Status_RS.Frg_RS_f_Schaeumen
   //    UN    "DB005_RS<->Extern".Status_RS.BA_Hand
   //    S     #St_Nr_053
   // 054Schäumroboter nicht in HP für Start Produktion
   //    U     "T_Start_RT_1"
   //    U     "DB151_Rundtisch_1".BA_Anlage.Automatik
   //    U     "DB005_RS<->Extern".Status_RS.Frg_Roboter_f_Schaeumen
   //    UN    "DB005_RS<->Extern".Status_RS.ABB_Schaeumen_HomePos
   //    UN    "DB005_RS<->Extern".Status_RS.BA_Hand
   //    S     #St_Nr_054
   // 055 Schäummaschine nicht bereit
   //    U     "T_Start_RT_1"
   //    U     "DB151_Rundtisch_1".BA_Anlage.Automatik
   //    UN    "DB005_RS<->Extern".Status_RS.Frg_RS_f_Schaeumen
   //    UN    "DB005_RS<->Extern".Status_RS.BA_Hand
   //    S     #St_Nr_055
   // 056 PT100 Vorlauf Wasser defekt
   //    U     "DB011_ZEITEN".RT_1_F_Sensor_Temp_VL
   //    S     #St_Nr_056
   // 057 PT100 Rücklauf Wasser defekt
   //    U     "DB011_ZEITEN".RT_1_F_Sensor_Temp_RL
   //    S     #St_Nr_057
   // 058 Max Warnung  Wassertemperatur
   //    U     "DB011_ZEITEN".RT_1_STG_Warn_Max
   //    S     #St_Nr_058
   // 059 Min Warnung Wassertemperatur
   //    U     "DB011_ZEITEN".RT_1_STG_Warn_Min
   //    S     #St_Nr_059
   // 060 Max Störung Wassertemperatur
   //    U     "DB011_ZEITEN".RT_1_STG_Tol_Max
   //    S     #St_Nr_060
   // 061 Min Störung Wassertemperatur
   //    U     "DB011_ZEITEN".RT_1_STG_Tol_Min
   //    S     #St_Nr_061
   // 062 Störung Versorgung Druckluft
   //    S     #St_Nr_062
   // 063 Nicht alle FTs gesteckt
   //    S     #St_Nr_063
   // 064 Sicherung Maschine
   //    S     #St_Nr_064
   // 065 Versorgung der Temperiergeräte
   //    S     #St_Nr_065
   // 066 Reserve
   //    S     #St_Nr_066
   // 067 Reserve
   //    S     #St_Nr_067
   // 068 Reserve
   //    S     #St_Nr_068
   // 069 Reserve
   //    S     #St_Nr_069
   // 070 Reserve
   //    S     #St_Nr_070
   // 071 Reserve
   //    S     #St_Nr_071
   // 072 Reserve
   //    S     #St_Nr_072
   // 073 Reserve
   //    S     #St_Nr_073
   // 074 Reserve
   //    S     #St_Nr_074
   // 075 Reserve
   //    S     #St_Nr_075
   // 076 Reseve
   //    S     #St_Nr_076
   // 077 Segment 01 ist nicht erreichbar
   //    S     #St_Nr_077
   // 078 Segment 02 ist nicht erreichbar
   //    S     #St_Nr_078
   // 079 Segment 03 ist nicht erreichbar
   //    S     #St_Nr_079
   // 080 Segment 04 ist nicht erreichbar
   //    S     #St_Nr_080
   // 081 Segment 05 ist nicht erreichbar
   //    S     #St_Nr_081
   // 082 Segment 06 ist nicht erreichbar
   //    S     #St_Nr_082
   // 083 Segment 07 ist nicht erreichbar
   //    S     #St_Nr_083
   // 084 Segment 08 ist nicht erreichbar
   //    S     #St_Nr_084
   // 085 Segment 09 ist nicht erreichbar
   //    S     #St_Nr_085
   // 086 Segment 10 ist nicht erreichbar
   //    S     #St_Nr_086
   // 08 7Segment 11 ist nicht erreichbar
   //      S     #St_Nr_087
   // 088 Segment 12 ist nicht erreichbar
   //      S     #St_Nr_088
   // 089 Segment 13 ist nicht erreichbar
   //       S     #St_Nr_089
   // 090 Segment 14 ist nicht erreichbar
   //       S     #St_Nr_090
   // 091 Segment 15 ist nicht erreichbar
   //      S     #St_Nr_091
   // 092 Segment 16 ist nicht erreichbar
   //      S     #St_Nr_092
   // 093 Segment 17 ist nicht erreichbar
   //      S     #St_Nr_093
   // 094 Segment 18 ist nicht erreichbar
   //      S     #St_Nr_094
   // 095 Segment 19 ist nicht erreichbar
   //      S     #St_Nr_095
   // 096 Segment 20 ist nicht erreichbar
   //      S     #St_Nr_096
END_REGION

REGION Network 5: Ablöschen der Meldungen
   // Die lokalen Variablen der Meldungen können immer abgelöscht werden, da diese in 
   // dem nachfolgendem Netzwerk immer neu zugewiesen werden. 
   // Würden die lokalen Variablen nicht gelöscht werden, könnte es vorkommen, daß 
   // eine auskommentierte Meldung nicht mehr zurückgesetzt werden könnte da diese im 
   // Datenbaustein noch gespeichert ist.
         L     12;  // Interner Offset für Meldungen
         SLD   3;
         LAR1;  // Adresse für lokale Meldungen
   //
         L     2;  // Anzahl der Meldungsworte
   M006: T     #Schleifenzaehler;  //
   //
         L     0;  // Lokale Meldungen zurücksetzten
         T     LW[AR1, P#0.0];  //
   //
         +AR1  P#2.0;
   //
         L     #Schleifenzaehler;  // Wenn Schleifenzähler <> 0
         LOOP  M006;  // Schleife erneut durchlaufen
END_REGION

REGION Network 6: Meldungen
         NOP   0;
   // 097: Not- Halt Taster am Schaltschrank wurde betätigt
   //    U
   //    =     "DB1010_Fault".ES.ControlCabinet
   //    =     #Mld_Nr_097
   // 098: Not- Halt- Taster am Bedienpult  betätigt
         A     "ES_TT_operating_panel";
         =     "DB1010_TT_Fault".ES.Operatingpanel;
         =     #Mld_Nr_098;
   // 099: Not- Halt- Taster 3  betätigt
   //    =     "DB1010_Fault".ES.Handling_2
   //    =     #Mld_Nr_099
   // 100: Not- Halt von der PU Maschine steht an
   //    UN    "ES_Machine"
   //    =     "DB1010_Fault".ES.ES_machine
   //    =     #Mld_Nr_100
   // 101: Taktdehnung ist aktiv
   //    =     #Mld_Nr_101
   // 102: Steuerspannung fehlt
         AN    "ES_TT_operating_panel";
         AN    "ES_foaming_machine";
         AN    "DB1001_TT_State".BA_Anlage.Steuerspannung_ein;
         =     #Mld_Nr_102;
   // 103: Vorwahl Schutztür WW ist aktiv
   //       U     "HM_Aw_Tuer_WW_Oeff_RT1"
   //       U     "E_Tuer_WW_ok_RT_1"
   //       =     #Mld_Nr_103
   // 104: Anlage stoppt für Teachen der Roboterbahn
         O     "DB1001_TT_State".Bits.Stop_fuer_Teachen;
         =     #Mld_Nr_104;
   // 105: Anlage stoppt für Werkzeugwechsel
         O     "DB1001_TT_State".Bits.Stop_fuer_WW;
         =     #Mld_Nr_105;
   // 106: NH Relais auf RT nicht quittiert
         AN    "DB1031_AddStatus".SaftyDevice[1].HFforMESAutomaticStop;
         AN    "DB1031_AddStatus".SaftyDevice[1].HFforMESAutomaticStop;
         AN    "DB1031_AddStatus".SaftyDevice[2].HFforMESAutomaticStop;
         AN    "DB1031_AddStatus".SaftyDevice[4].HFforMESAutomaticStop;
         A     "AS_pendelum_flap_to_handling";
         A     "AS_pendelum_flap_from_handling";
         AN    "DB1001_TT_State".BA_Anlage.Automatik_Stop_ok;
         A     "DB1001_TT_State".BA_Anlage.Steuerspannung_ein;
         =     #Mld_Nr_106;
   // 107: NH von PU
   //    =     #Mld_Nr_107
   // 108: NA Roboter
   //       U     "NA_Roboter"
   //       =     #Mld_Nr_108
   // 109: WZW Tür nicht geschlossen und quittiert
   //    =     #Mld_Nr_109
   // 110: Tür Roboter 1
   //      UN    "Tuer_2_quittiert"
   //      =     #Mld_Nr_110
   // 111: Tür Roboter 2 (Trennen)
   //      UN    "Tuer_3_quittiert"
   //      =     #Mld_Nr_111
   // 112: Pendelklappe 1
         AN    "AS_pendelum_flap_to_handling";
         =     #Mld_Nr_112;
   // 113: Pendelklappe 2
         AN    "AS_pendelum_flap_from_handling";
         =     #Mld_Nr_113;
   // -----------------------
         ON    "AS_pendelum_flap_to_handling";
         ON    "AS_pendelum_flap_from_handling";
         =     "DB1010_TT_Fault".AS.AS_WingDoor;
   // 114: Pendelklappe 3
   //    =     #Mld_Nr_114
   // 115: Pendelklappe 4
   //    =     #Mld_Nr_115
   // 116: NA Handling1
   //    =     #Mld_Nr_116
   // 117: NA Handling2
   //    =     #Mld_Nr_117
   // 118:NA Handling3
   //    =     #Mld_Nr_118
   // 119: Segment x wurde referenziert
         A     "DB1001_TT_State".IPOS.Status.BA_Referenzieren;
         =     #Mld_Nr_119;
   // 120: STG Relais Pendelklappe
   //    =     #Mld_Nr_120
   // 121: Reserve
   //    =     #Mld_Nr_121
   // 122: Drehsperre von RT2 wegen Teachen angewählt
   //      U     "DB152_Rundtisch_2".Bits.Stop_fuer_Teachen
   //      =     #Mld_Nr_122
   // 123: Drehsperre von IRB 1
   //      U     "DB005_RS<->Extern".Status_RS.ABB_Schaeumen_Drehsperre
   //      L     S5T#1M
   //      SE    T     57
   //      U     T     57
   //      =     #Mld_Nr_123
   // 124: Drehsperre von IRB 2
   //      UN    "DB051_KUKA".Status_Roboter_KUKA.Input_vom_Roboter.E_KRC_OUT_ausserhalb
   //      L     S5T#1M
   //      SE    T     58
   //      U     T     58
   //      =     #Mld_Nr_124

   // 125: Rundtisch nicht in Position SEW
         A     "DB1001_TT_State".BA_Anlage.Start_Produktion;
         AN    "DB1001_TT_State".IPOS.Status.RT_in_Position;
         A     "DB1001_TT_State".IPOS.Status.IPOS_referenziert;
         AN    "DB1001_TT_State".IPOS.Status.RT_dreht;
         =     #Mld_Nr_125;
   // 126: Der Rundtisch ist noch nicht referenziert
         AN    "DB1001_TT_State".IPOS.Status.IPOS_referenziert;
         =     #Mld_Nr_126;
   // 127: Funktion "Leerfahren" des Rundtisches ist angewählt
   //      U     "DB1001_RT".Status.S_RT_Leerfahren
   //      UN    "DB1001_RT".Status.RT_ist_leergefahren
   //      =     #Mld_Nr_127
   // 128: Alle Werkzeuge sind in Abwahlposition oder nicht Freigegeben
   //      U     "DB_RT<->Extern".Status_RT_1.RT_ist_leergefahren
   //      =     #Mld_Nr_128
END_REGION

REGION Network 7: Störungsgruppe 1 und Änderung ermitteln; Bits -> DB für Anzeige
         L     0;  // Interner Offset für Störungsgruppe 1
         SLD   3;  //
         LAR1;  // Adresse für lokale Störungen
   //
         L     0;  // Interner Offset für Störungsgruppe 1
         L     #IN_Start_Stoerungen;
         +D;
         SLD   3;  //
         LAR2;  // Adresse für Störung im DB
   //
         L     2;  // Anzahl der Störungsworte
   M003: T     #Schleifenzaehler;  //
   //
         OPN   #IN_DB_Stoerungen;  //
         L     DBW[AR2, P#0.0];  // Gespeicherte Störung mit
         L     LW[AR1, P#0.0];  // Lokale Störung       vergleichen
         <>D;  //
         T     DBW[AR2, P#0.0];  // im DB speichern und
         S     #IO_Daten_Senden;  // Sendeanforderung an PU (FB120)
         S     #IO_Stoerungsaenderung;  // Störungsanderung für Störauswertung (FB9)
         S     #IO_Stoer_Grp_1_aktiv;  // und Sammelsignal setzen
   //
         +AR1  P#2.0;
         +AR2  P#2.0;
   //
         L     #Schleifenzaehler;  // Wenn Schleifenzähler <> 0
         LOOP  M003;  // Schleife erneut durchlaufen
   //
         A     #IN_Stoer_Grp_1_von_Ext;  // Storung vom Rechner
         AN    #IN_Reset_fault_Grp;  // in die SPS einbinden
         FP    #IO_FM_Stoer_Grp_1_v_Ext;
         S     #IO_Stoerungsaenderung;
         S     #IO_Stoer_Grp_1_aktiv;
END_REGION
